// TIA Portal project "OC_test_FFT" (V13)

(* hardware
DEVICE "OpenController"  CPU 1515SP PC
   slot 0: "OpenController"  CPU 1515SP PC  6ES7 677-2AAxx-0xB0  V1.8
      slot 124: "Diagbase"  Diagbase  V6.0.4
      slot 125: "OpenController"  PC Station 2.0  Station_Manager  V2.0
   slot 1: "CPU1505S"  CPU 1505S  6ES7 672-5AC00-0YA0  V1.8
   slot 2: "PROFINET onboard_2"  IE General  IE_CP  V2.0
   slot 4: "HMI_RT_1"  WinCC RT Advanced  6AV2 104-0xxxx-xxxx  13.0.1.0
      slot 33792: "Host interface"  Host interface
   slot 127: "PROFINET BusAdapter CU"  PROFINET Interface  6ES7 193-6AR00-0AA0  V0.0
      slot 32769: "Port_1"  6ES7 193-6AR00-0AA0
      slot 32770: "Port_2"  6ES7 193-6AR00-0AA0
   slot 1002: "Server module_1"  Server module  6ES7 193-6PA00-0AA0  V1.0
      slot 1: "Server module_1"  Server module  6ES7 193-6PA00-0AA0
*)

// ===== PLC "CPU1505S"  CPU 1505S =====

VAR_GLOBAL   // PLC tag table "Default tag table"
   "System_Byte" AT %MB1 : Byte;
   "FirstScan" AT %M1.0 : Bool;
   "DiagStatusUpdate" AT %M1.1 : Bool;
   "AlwaysTRUE" AT %M1.2 : Bool;
   "AlwaysFALSE" AT %M1.3 : Bool;
   "Clock_Byte" AT %MB0 : Byte;
   "Clock_10Hz" AT %M0.0 : Bool;
   "Clock_5Hz" AT %M0.1 : Bool;
   "Clock_2.5Hz" AT %M0.2 : Bool;
   "Clock_2Hz" AT %M0.3 : Bool;
   "Clock_1.25Hz" AT %M0.4 : Bool;
   "Clock_1Hz" AT %M0.5 : Bool;
   "Clock_0.625Hz" AT %M0.6 : Bool;
   "Clock_0.5Hz" AT %M0.7 : Bool;
END_VAR

TYPE "FFT_Filter_RTComplex"
   STRUCT
      re : Real;
      im : Real;
   END_STRUCT;
END_TYPE

DATA_BLOCK "ODK_Params"   // DB1
{ S7_Optimized_Access := 'FALSE' }
VERSION : 0.1
   VAR
      Filter_Load : Struct
      END_STRUCT;
      Filt1 : Struct
      END_STRUCT;
      Filt2 : Struct
      END_STRUCT;
      WaveInput_Load : Struct
      END_STRUCT;
      WaveSetup : Struct
      END_STRUCT;
      GetSamples : Struct
      END_STRUCT;
      WriteSamples : Struct
      END_STRUCT;
   END_VAR
BEGIN
END_DATA_BLOCK

DATA_BLOCK "FFT_Filter_RT_Load_DB"   // DB2
{ S7_Optimized_Access := 'FALSE' }
VERSION : 0.1
// stored: InstanceOfName FFT_Filter_RT_Load
"FFT_Filter_RT_Load"
BEGIN
END_DATA_BLOCK

DATA_BLOCK "FFT_Filter_RTFFT_Filt_DB"   // DB3
{ S7_Optimized_Access := 'FALSE' }
VERSION : 0.1
// stored: InstanceOfName FFT_Filter_RTFFT_Filt
"FFT_Filter_RTFFT_Filt"
BEGIN
END_DATA_BLOCK

DATA_BLOCK "FFT_Filter_RTFFT_Filt_DB_1"   // DB4
{ S7_Optimized_Access := 'FALSE' }
VERSION : 0.1
// stored: InstanceOfName FFT_Filter_RTFFT_Filt
"FFT_Filter_RTFFT_Filt"
BEGIN
END_DATA_BLOCK

DATA_BLOCK "FFT_Filt_Data_Load_DB"   // DB5
{ S7_Optimized_Access := 'FALSE' }
VERSION : 0.1
// stored: InstanceOfName FFT_Filt_Data_Load
"FFT_Filt_Data_Load"
BEGIN
END_DATA_BLOCK

DATA_BLOCK "FFT_Filt_DataWaveSetup_DB"   // DB6
{ S7_Optimized_Access := 'FALSE' }
VERSION : 0.1
// stored: InstanceOfName FFT_Filt_DataWaveSetup
"FFT_Filt_DataWaveSetup"
BEGIN
END_DATA_BLOCK

DATA_BLOCK "FFT_Filt_DataGetSamplesStereo_DB"   // DB7
{ S7_Optimized_Access := 'FALSE' }
VERSION : 0.1
// stored: InstanceOfName FFT_Filt_DataGetSamplesStereo
"FFT_Filt_DataGetSamplesStereo"
BEGIN
END_DATA_BLOCK

DATA_BLOCK "FFT_Filt_DataWriteSamples_DB"   // DB8
{ S7_Optimized_Access := 'FALSE' }
VERSION : 0.1
// stored: InstanceOfName FFT_Filt_DataWriteSamples
"FFT_Filt_DataWriteSamples"
BEGIN
END_DATA_BLOCK

FUNCTION_BLOCK "FFT_Filter_RT_Load"   // FB1, SCL
{ S7_Optimized_Access := 'FALSE' }
VERSION : 0.1
// This block is AUTO GENERATED - DO NOT MODIFY this block!
// Created by ODK_CodeGenerator version 2.0.0.0
// at Sun January 31 20:03:01 2016
// ********************************************************
BEGIN
   //
   // DO NOT CHANGE BELOW OF THIS LINE !!
   // This is an automatic generated block by the
   // ODK_CodeGenerator version 2.0.0.0
   // DO NOT CHANGE !!
   //
   #ODK_Load_Instance(REQ := #REQ,
                      LIBRARY_NAME := #_odk_internal_LIBRARY_NAME,
                      INSTANCE_ID := #_odk_internal_INSTANCE_ID,
                      DONE => #DONE,
                      BUSY => #BUSY,
                      ERROR => #ERROR,
                      STATUS => #STATUS);
   //
   // DO NOT CHANGE !!
   // This is an automatic generated block by the
   // ODK_CodeGenerator version 2.0.0.0
   // DO NOT CHANGE ABOVE OF THIS LINE !!
   //
END_FUNCTION_BLOCK

FUNCTION_BLOCK "FFT_Filter_RT_Unload"   // FB2, SCL
{ S7_Optimized_Access := 'FALSE' }
VERSION : 0.1
// This block is AUTO GENERATED - DO NOT MODIFY this block!
// Created by ODK_CodeGenerator version 2.0.0.0
// at Sun January 31 20:03:01 2016
// ********************************************************
BEGIN
   //
   // DO NOT CHANGE BELOW OF THIS LINE !!
   // This is an automatic generated block by the
   // ODK_CodeGenerator version 2.0.0.0
   // DO NOT CHANGE !!
   //
   #ODK_Unld_Instance(REQ := #REQ,
                      INSTANCE_ID := #_odk_internal_INSTANCE_ID,
                      DONE => #DONE,
                      BUSY => #BUSY,
                      ERROR => #ERROR,
                      STATUS => #STATUS);
   //
   // DO NOT CHANGE !!
   // This is an automatic generated block by the
   // ODK_CodeGenerator version 2.0.0.0
   // DO NOT CHANGE ABOVE OF THIS LINE !!
   //
END_FUNCTION_BLOCK

FUNCTION_BLOCK "FFT_Filter_RTFFT1024p"   // FB3, SCL
{ S7_Optimized_Access := 'FALSE' }
VERSION : 0.1
// This block is AUTO GENERATED - DO NOT MODIFY this block!
// Created by ODK_CodeGenerator version 2.0.0.0
// at Sun January 31 20:03:01 2016
// ********************************************************
BEGIN
   //
   // DO NOT CHANGE BELOW OF THIS LINE !!
   // This is an automatic generated block by the
   // ODK_CodeGenerator version 2.0.0.0
   // DO NOT CHANGE !!
   //
   #_odk_internal_pos := 0;
   FOR #_odk_internal_i := 0 TO 1023 DO
     #_odk_internal_err := WRITE_LITTLE(src_variable := #timeCoef[#_odk_internal_i], dest_array := #_odk_internal_IN_BUFFER, pos := #_odk_internal_pos);
   END_FOR;
   #STATUS := ODK_ExcS(INSTANCE_ID := #_odk_internal_INSTANCE_ID,
                       COMMAND := #_odk_internal_COMMAND,
                       IN_DATA := #_odk_internal_IN_BUFFER,
                       INOUT_DATA := #_odk_internal_tmpDefaultValue,
                       OUT_DATA := #_odk_internal_OUT_BUFFER
   );
   IF #STATUS < 16#7000 THEN
     #_odk_internal_pos := 0;
     FOR #_odk_internal_udt_0 := 0 TO 1023 DO
       #_odk_internal_err := READ_LITTLE(dest_Variable => #freqCoef[#_odk_internal_udt_0].re, src_array := #_odk_internal_OUT_BUFFER, pos := #_odk_internal_pos);
       #_odk_internal_err := READ_LITTLE(dest_Variable => #freqCoef[#_odk_internal_udt_0].im, src_array := #_odk_internal_OUT_BUFFER, pos := #_odk_internal_pos);
     END_FOR;
   END_IF;
   //
   // DO NOT CHANGE !!
   // This is an automatic generated block by the
   // ODK_CodeGenerator version 2.0.0.0
   // DO NOT CHANGE ABOVE OF THIS LINE !!
   //
END_FUNCTION_BLOCK

FUNCTION_BLOCK "FFT_Filter_RTLP_Filter"   // FB4, SCL
{ S7_Optimized_Access := 'FALSE' }
VERSION : 0.1
// This block is AUTO GENERATED - DO NOT MODIFY this block!
// Created by ODK_CodeGenerator version 2.0.0.0
// at Sun January 31 20:03:01 2016
// ********************************************************
BEGIN
   //
   // DO NOT CHANGE BELOW OF THIS LINE !!
   // This is an automatic generated block by the
   // ODK_CodeGenerator version 2.0.0.0
   // DO NOT CHANGE !!
   //
   #_odk_internal_pos := 0;
   FOR #_odk_internal_udt_0 := 0 TO 1023 DO
     #_odk_internal_err := WRITE_LITTLE(src_variable := #freqCoef[#_odk_internal_udt_0].re, dest_array := #_odk_internal_IN_BUFFER, pos := #_odk_internal_pos);
     #_odk_internal_err := WRITE_LITTLE(src_variable := #freqCoef[#_odk_internal_udt_0].im, dest_array := #_odk_internal_IN_BUFFER, pos := #_odk_internal_pos);
   END_FOR;
   #STATUS := ODK_ExcS(INSTANCE_ID := #_odk_internal_INSTANCE_ID,
                       COMMAND := #_odk_internal_COMMAND,
                       IN_DATA := #_odk_internal_IN_BUFFER,
                       INOUT_DATA := #_odk_internal_tmpDefaultValue,
                       OUT_DATA := #_odk_internal_OUT_BUFFER
   );
   IF #STATUS < 16#7000 THEN
     #_odk_internal_pos := 0;
     FOR #_odk_internal_udt_0 := 0 TO 1023 DO
       #_odk_internal_err := READ_LITTLE(dest_Variable => #freqCoefFilt[#_odk_internal_udt_0].re, src_array := #_odk_internal_OUT_BUFFER, pos := #_odk_internal_pos);
       #_odk_internal_err := READ_LITTLE(dest_Variable => #freqCoefFilt[#_odk_internal_udt_0].im, src_array := #_odk_internal_OUT_BUFFER, pos := #_odk_internal_pos);
     END_FOR;
   END_IF;
   //
   // DO NOT CHANGE !!
   // This is an automatic generated block by the
   // ODK_CodeGenerator version 2.0.0.0
   // DO NOT CHANGE ABOVE OF THIS LINE !!
   //
END_FUNCTION_BLOCK

FUNCTION_BLOCK "FFT_Filter_RTIFFT1024p"   // FB5, SCL
{ S7_Optimized_Access := 'FALSE' }
VERSION : 0.1
// This block is AUTO GENERATED - DO NOT MODIFY this block!
// Created by ODK_CodeGenerator version 2.0.0.0
// at Sun January 31 20:03:01 2016
// ********************************************************
BEGIN
   //
   // DO NOT CHANGE BELOW OF THIS LINE !!
   // This is an automatic generated block by the
   // ODK_CodeGenerator version 2.0.0.0
   // DO NOT CHANGE !!
   //
   #_odk_internal_pos := 0;
   FOR #_odk_internal_udt_0 := 0 TO 1023 DO
     #_odk_internal_err := WRITE_LITTLE(src_variable := #freqCoef[#_odk_internal_udt_0].re, dest_array := #_odk_internal_IN_BUFFER, pos := #_odk_internal_pos);
     #_odk_internal_err := WRITE_LITTLE(src_variable := #freqCoef[#_odk_internal_udt_0].im, dest_array := #_odk_internal_IN_BUFFER, pos := #_odk_internal_pos);
   END_FOR;
   #STATUS := ODK_ExcS(INSTANCE_ID := #_odk_internal_INSTANCE_ID,
                       COMMAND := #_odk_internal_COMMAND,
                       IN_DATA := #_odk_internal_IN_BUFFER,
                       INOUT_DATA := #_odk_internal_tmpDefaultValue,
                       OUT_DATA := #_odk_internal_OUT_BUFFER
   );
   IF #STATUS < 16#7000 THEN
     #_odk_internal_pos := 0;
     FOR #_odk_internal_i := 0 TO 1023 DO
       #_odk_internal_err := READ_LITTLE(dest_Variable => #timeCoefOut[#_odk_internal_i], src_array := #_odk_internal_OUT_BUFFER, pos := #_odk_internal_pos);
     END_FOR;
   END_IF;
   //
   // DO NOT CHANGE !!
   // This is an automatic generated block by the
   // ODK_CodeGenerator version 2.0.0.0
   // DO NOT CHANGE ABOVE OF THIS LINE !!
   //
END_FUNCTION_BLOCK

FUNCTION_BLOCK "FFT_Filter_RTFFT_Filt"   // FB6, SCL
{ S7_Optimized_Access := 'FALSE' }
VERSION : 0.1
// This block is AUTO GENERATED - DO NOT MODIFY this block!
// Created by ODK_CodeGenerator version 2.0.0.0
// at Sun January 31 20:03:01 2016
// ********************************************************
BEGIN
   //
   // DO NOT CHANGE BELOW OF THIS LINE !!
   // This is an automatic generated block by the
   // ODK_CodeGenerator version 2.0.0.0
   // DO NOT CHANGE !!
   //
   #_odk_internal_pos := 0;
   FOR #_odk_internal_i := 0 TO 1023 DO
     #_odk_internal_err := WRITE_LITTLE(src_variable := #timeCoef[#_odk_internal_i], dest_array := #_odk_internal_IN_BUFFER, pos := #_odk_internal_pos);
   END_FOR;
   #STATUS := ODK_ExcS(INSTANCE_ID := #_odk_internal_INSTANCE_ID,
                       COMMAND := #_odk_internal_COMMAND,
                       IN_DATA := #_odk_internal_IN_BUFFER,
                       INOUT_DATA := #_odk_internal_tmpDefaultValue,
                       OUT_DATA := #_odk_internal_OUT_BUFFER
   );
   IF #STATUS < 16#7000 THEN
     #_odk_internal_pos := 0;
     FOR #_odk_internal_i := 0 TO 1023 DO
       #_odk_internal_err := READ_LITTLE(dest_Variable => #timeCoefOut[#_odk_internal_i], src_array := #_odk_internal_OUT_BUFFER, pos := #_odk_internal_pos);
     END_FOR;
   END_IF;
   //
   // DO NOT CHANGE !!
   // This is an automatic generated block by the
   // ODK_CodeGenerator version 2.0.0.0
   // DO NOT CHANGE ABOVE OF THIS LINE !!
   //
END_FUNCTION_BLOCK

FUNCTION_BLOCK "FFT_Filt_Data_Load"   // FB7, SCL
{ S7_Optimized_Access := 'FALSE' }
VERSION : 0.1
// This block is AUTO GENERATED - DO NOT MODIFY this block!
// Created by ODK_CodeGenerator version 2.0.0.0
// at Sun January 17 17:54:04 2016
// ********************************************************
BEGIN
   //
   // DO NOT CHANGE BELOW OF THIS LINE !!
   // This is an automatic generated block by the
   // ODK_CodeGenerator version 2.0.0.0
   // DO NOT CHANGE !!
   //
   #ODK_Load_Instance(REQ := #REQ,
                      LIBRARY_NAME := #_odk_internal_LIBRARY_NAME,
                      INSTANCE_ID := #_odk_internal_INSTANCE_ID,
                      DONE => #DONE,
                      BUSY => #BUSY,
                      ERROR => #ERROR,
                      STATUS => #STATUS);
   //
   // DO NOT CHANGE !!
   // This is an automatic generated block by the
   // ODK_CodeGenerator version 2.0.0.0
   // DO NOT CHANGE ABOVE OF THIS LINE !!
   //
END_FUNCTION_BLOCK

FUNCTION_BLOCK "FFT_Filt_Data_Unload"   // FB8, SCL
{ S7_Optimized_Access := 'FALSE' }
VERSION : 0.1
// This block is AUTO GENERATED - DO NOT MODIFY this block!
// Created by ODK_CodeGenerator version 2.0.0.0
// at Sun January 17 17:54:04 2016
// ********************************************************
BEGIN
   //
   // DO NOT CHANGE BELOW OF THIS LINE !!
   // This is an automatic generated block by the
   // ODK_CodeGenerator version 2.0.0.0
   // DO NOT CHANGE !!
   //
   #ODK_Unld_Instance(REQ := #REQ,
                      INSTANCE_ID := #_odk_internal_INSTANCE_ID,
                      DONE => #DONE,
                      BUSY => #BUSY,
                      ERROR => #ERROR,
                      STATUS => #STATUS);
   //
   // DO NOT CHANGE !!
   // This is an automatic generated block by the
   // ODK_CodeGenerator version 2.0.0.0
   // DO NOT CHANGE ABOVE OF THIS LINE !!
   //
END_FUNCTION_BLOCK

FUNCTION_BLOCK "FFT_Filt_DataWaveSetup"   // FB9, SCL
{ S7_Optimized_Access := 'FALSE' }
VERSION : 0.1
// This block is AUTO GENERATED - DO NOT MODIFY this block!
// Created by ODK_CodeGenerator version 2.0.0.0
// at Sun January 17 17:54:04 2016
// ********************************************************
//  Setup file handles for IO operation
BEGIN
   //
   // DO NOT CHANGE BELOW OF THIS LINE !!
   // This is an automatic generated block by the
   // ODK_CodeGenerator version 2.0.0.0
   // DO NOT CHANGE !!
   //
   // Setup file handles for IO operation
   IF NOT #_odk_internal_Last_REQ & #REQ & NOT #BUSY THEN
     #_odk_internal_pos := 0;
     #_odk_internal_tmpStringLen := INT_TO_BYTE(LEN(#inFileName));
     #_odk_internal_IN_BUFFER[#_odk_internal_pos] := BYTE#254;
     #_odk_internal_pos := #_odk_internal_pos + 1;
     #_odk_internal_IN_BUFFER[#_odk_internal_pos] := #_odk_internal_tmpStringLen;
     #_odk_internal_pos := #_odk_internal_pos + 1;
     FOR #_odk_internal_i := 1 TO BYTE_TO_INT(#_odk_internal_tmpStringLen) DO
       #_odk_internal_IN_BUFFER[#_odk_internal_pos] := CHAR_TO_BYTE(#inFileName[#_odk_internal_i]);
       #_odk_internal_pos := #_odk_internal_pos + 1;
     END_FOR;
     #_odk_internal_pos := #_odk_internal_pos + 254 - #_odk_internal_tmpStringLen;
     #_odk_internal_tmpStringLen := INT_TO_BYTE(LEN(#outFileName));
     #_odk_internal_IN_BUFFER[#_odk_internal_pos] := BYTE#254;
     #_odk_internal_pos := #_odk_internal_pos + 1;
     #_odk_internal_IN_BUFFER[#_odk_internal_pos] := #_odk_internal_tmpStringLen;
     #_odk_internal_pos := #_odk_internal_pos + 1;
     FOR #_odk_internal_i := 1 TO BYTE_TO_INT(#_odk_internal_tmpStringLen) DO
       #_odk_internal_IN_BUFFER[#_odk_internal_pos] := CHAR_TO_BYTE(#outFileName[#_odk_internal_i]);
       #_odk_internal_pos := #_odk_internal_pos + 1;
     END_FOR;
     #_odk_internal_pos := #_odk_internal_pos + 254 - #_odk_internal_tmpStringLen;

   END_IF;
   #_odk_internal_Last_REQ := #REQ;
   #ODK_ExcA_Instance(REQ := #REQ,
                      INSTANCE_ID := #_odk_internal_INSTANCE_ID,
                      COMMAND := #_odk_internal_COMMAND,
                      IN_DATA := #_odk_internal_IN_BUFFER,
                      INOUT_DATA := #_odk_internal_tmpDefaultValue,
                      OUT_DATA := #_odk_internal_tmpDefaultValue,
                      DONE => #DONE,
                      BUSY => #BUSY,
                      ERROR => #ERROR,
                      STATUS => #STATUS);
   //
   // DO NOT CHANGE !!
   // This is an automatic generated block by the
   // ODK_CodeGenerator version 2.0.0.0
   // DO NOT CHANGE ABOVE OF THIS LINE !!
   //
END_FUNCTION_BLOCK

FUNCTION_BLOCK "FFT_Filt_DataGetSamplesStereo"   // FB10, SCL
{ S7_Optimized_Access := 'FALSE' }
VERSION : 0.1
// This block is AUTO GENERATED - DO NOT MODIFY this block!
// Created by ODK_CodeGenerator version 2.0.0.0
// at Sun January 17 17:54:04 2016
// ********************************************************
//  Get one filter samlple for processing
BEGIN
   //
   // DO NOT CHANGE BELOW OF THIS LINE !!
   // This is an automatic generated block by the
   // ODK_CodeGenerator version 2.0.0.0
   // DO NOT CHANGE !!
   //
   // Get one filter samlple for processing   
   #_odk_internal_Last_REQ := #REQ;
   #ODK_ExcA_Instance(REQ := #REQ,
                      INSTANCE_ID := #_odk_internal_INSTANCE_ID,
                      COMMAND := #_odk_internal_COMMAND,
                      IN_DATA := #_odk_internal_tmpDefaultValue,
                      INOUT_DATA := #_odk_internal_tmpDefaultValue,
                      OUT_DATA := #_odk_internal_OUT_BUFFER,
                      DONE => #DONE,
                      BUSY => #BUSY,
                      ERROR => #ERROR,
                      STATUS => #STATUS);
   IF NOT #BUSY & #_odk_internal_Last_BUSY & NOT #ERROR THEN
     #_odk_internal_pos := 0;
     FOR #_odk_internal_i := 0 TO 1023 DO
       #_odk_internal_err := READ_LITTLE(dest_Variable => #inputSamplesL[#_odk_internal_i], src_array := #_odk_internal_OUT_BUFFER, pos := #_odk_internal_pos);
     END_FOR;
     FOR #_odk_internal_i := 0 TO 1023 DO
       #_odk_internal_err := READ_LITTLE(dest_Variable => #inputSamplesR[#_odk_internal_i], src_array := #_odk_internal_OUT_BUFFER, pos := #_odk_internal_pos);
     END_FOR;
     #lastSample := BYTE_TO_BOOL(#_odk_internal_OUT_BUFFER[#_odk_internal_pos]);
     #_odk_internal_pos := #_odk_internal_pos + 1;
   END_IF;
   #_odk_internal_Last_BUSY := #BUSY;
   //
   // DO NOT CHANGE !!
   // This is an automatic generated block by the
   // ODK_CodeGenerator version 2.0.0.0
   // DO NOT CHANGE ABOVE OF THIS LINE !!
   //
END_FUNCTION_BLOCK

FUNCTION_BLOCK "FFT_Filt_DataWriteSamples"   // FB11, SCL
{ S7_Optimized_Access := 'FALSE' }
VERSION : 0.1
// This block is AUTO GENERATED - DO NOT MODIFY this block!
// Created by ODK_CodeGenerator version 2.0.0.0
// at Sun January 17 17:54:04 2016
// ********************************************************
//  write processed sample frame into file
BEGIN
   //
   // DO NOT CHANGE BELOW OF THIS LINE !!
   // This is an automatic generated block by the
   // ODK_CodeGenerator version 2.0.0.0
   // DO NOT CHANGE !!
   //
   // write processed sample frame into file
   IF NOT #_odk_internal_Last_REQ & #REQ & NOT #BUSY THEN
     #_odk_internal_pos := 0;
     FOR #_odk_internal_i := 0 TO 1023 DO
       #_odk_internal_err := WRITE_LITTLE(src_variable := #filteredSamplesL[#_odk_internal_i], dest_array := #_odk_internal_IN_BUFFER, pos := #_odk_internal_pos);
     END_FOR;
     FOR #_odk_internal_i := 0 TO 1023 DO
       #_odk_internal_err := WRITE_LITTLE(src_variable := #filteredSamplesR[#_odk_internal_i], dest_array := #_odk_internal_IN_BUFFER, pos := #_odk_internal_pos);
     END_FOR;

   END_IF;
   #_odk_internal_Last_REQ := #REQ;
   #ODK_ExcA_Instance(REQ := #REQ,
                      INSTANCE_ID := #_odk_internal_INSTANCE_ID,
                      COMMAND := #_odk_internal_COMMAND,
                      IN_DATA := #_odk_internal_IN_BUFFER,
                      INOUT_DATA := #_odk_internal_tmpDefaultValue,
                      OUT_DATA := #_odk_internal_tmpDefaultValue,
                      DONE => #DONE,
                      BUSY => #BUSY,
                      ERROR => #ERROR,
                      STATUS => #STATUS);
   //
   // DO NOT CHANGE !!
   // This is an automatic generated block by the
   // ODK_CodeGenerator version 2.0.0.0
   // DO NOT CHANGE ABOVE OF THIS LINE !!
   //
END_FUNCTION_BLOCK

FUNCTION "Filter_Run" : Void   // FC1, FBD
{ S7_Optimized_Access := 'FALSE' }
VERSION : 0.1
BEGIN

REGION Network 1
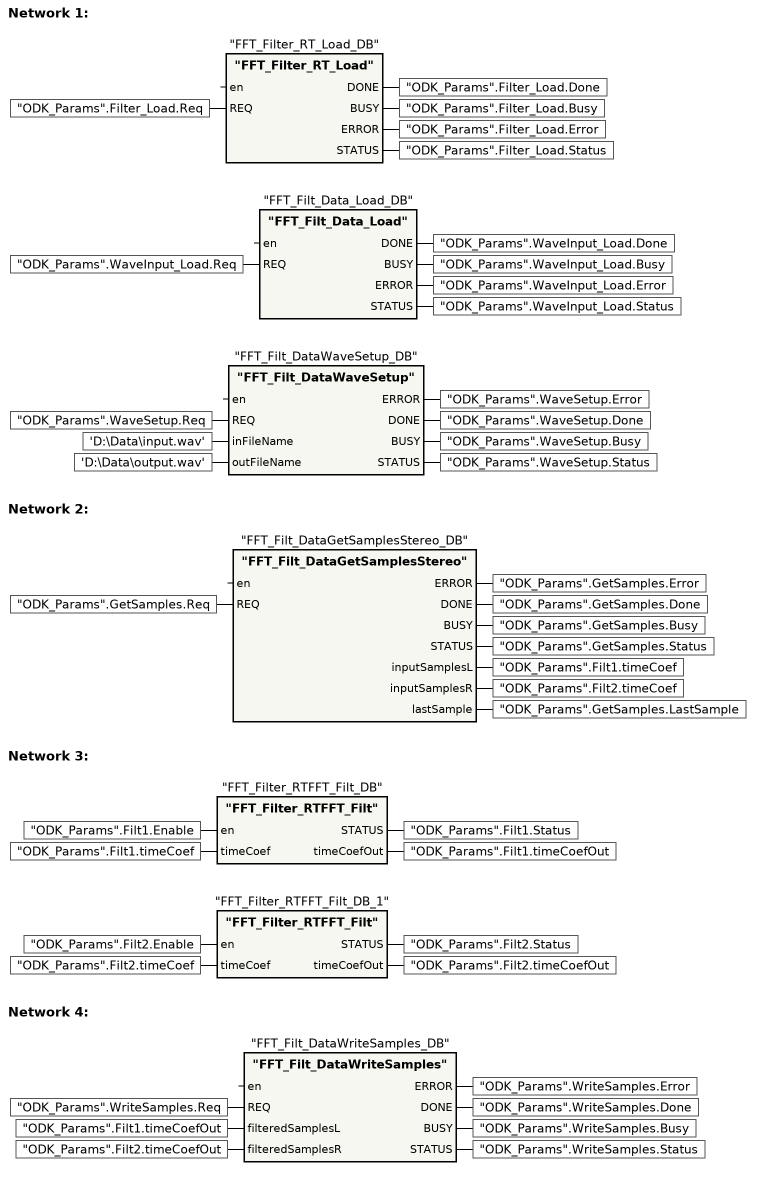
   "FFT_Filter_RT_Load_DB"(REQ := "ODK_Params".Filter_Load.Req,   // "FFT_Filter_RT_Load"
                           DONE => "ODK_Params".Filter_Load.Done,
                           BUSY => "ODK_Params".Filter_Load.Busy,
                           ERROR => "ODK_Params".Filter_Load.Error,
                           STATUS => "ODK_Params".Filter_Load.Status);
   "FFT_Filt_Data_Load_DB"(REQ := "ODK_Params".WaveInput_Load.Req,   // "FFT_Filt_Data_Load"
                           DONE => "ODK_Params".WaveInput_Load.Done,
                           BUSY => "ODK_Params".WaveInput_Load.Busy,
                           ERROR => "ODK_Params".WaveInput_Load.Error,
                           STATUS => "ODK_Params".WaveInput_Load.Status);
   "FFT_Filt_DataWaveSetup_DB"(REQ := "ODK_Params".WaveSetup.Req,   // "FFT_Filt_DataWaveSetup"
                           inFileName := 'D:\Data\input.wav',
                           outFileName := 'D:\Data\output.wav',
                           ERROR => "ODK_Params".WaveSetup.Error,
                           DONE => "ODK_Params".WaveSetup.Done,
                           BUSY => "ODK_Params".WaveSetup.Busy,
                           STATUS => "ODK_Params".WaveSetup.Status);
END_REGION

REGION Network 2
   "FFT_Filt_DataGetSamplesStereo_DB"(REQ := "ODK_Params".GetSamples.Req,   // "FFT_Filt_DataGetSamplesStereo"
                           ERROR => "ODK_Params".GetSamples.Error,
                           DONE => "ODK_Params".GetSamples.Done,
                           BUSY => "ODK_Params".GetSamples.Busy,
                           STATUS => "ODK_Params".GetSamples.Status,
                           inputSamplesL => "ODK_Params".Filt1.timeCoef,
                           inputSamplesR => "ODK_Params".Filt2.timeCoef,
                           lastSample => "ODK_Params".GetSamples.LastSample);
END_REGION

REGION Network 3
   IF "ODK_Params".Filt1.Enable THEN
       "FFT_Filter_RTFFT_Filt_DB"(timeCoef := "ODK_Params".Filt1.timeCoef,   // "FFT_Filter_RTFFT_Filt"
                               STATUS => "ODK_Params".Filt1.Status,
                               timeCoefOut => "ODK_Params".Filt1.timeCoefOut);
   END_IF;
   IF "ODK_Params".Filt2.Enable THEN
       "FFT_Filter_RTFFT_Filt_DB_1"(timeCoef := "ODK_Params".Filt2.timeCoef,   // "FFT_Filter_RTFFT_Filt"
                               STATUS => "ODK_Params".Filt2.Status,
                               timeCoefOut => "ODK_Params".Filt2.timeCoefOut);
   END_IF;
END_REGION

REGION Network 4
   "FFT_Filt_DataWriteSamples_DB"(REQ := "ODK_Params".WriteSamples.Req,   // "FFT_Filt_DataWriteSamples"
                           filteredSamplesL := "ODK_Params".Filt1.timeCoefOut,
                           filteredSamplesR := "ODK_Params".Filt2.timeCoefOut,
                           ERROR => "ODK_Params".WriteSamples.Error,
                           DONE => "ODK_Params".WriteSamples.Done,
                           BUSY => "ODK_Params".WriteSamples.Busy,
                           STATUS => "ODK_Params".WriteSamples.Status);
END_REGION
END_FUNCTION

ORGANIZATION_BLOCK "Main"   // OB1, LAD, ProgramCycle
TITLE = "Main Program Sweep (Cycle)"
{ S7_Optimized_Access := 'FALSE' }
VERSION : 0.1
BEGIN

REGION Network 1
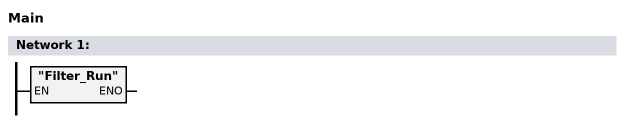
   RUNG wire#powerrail
      "Filter_Run"()
   END_RUNG
   // the same network as SCL:
   "Filter_Run"();
END_REGION
END_ORGANIZATION_BLOCK

(* ===== HMI "HMI_RT_1" =====
connection "HMI_Connection_1": Softbus, S7_1500_OMS

HMI tags "Default tag table"
   "ODK_Params_Filter_Load_Status" : Int, 100 ms
   "ODK_Params_Filter_Load_Req" : Bool, 100 ms
   "ODK_Params_WaveInput_Load_Status" : Int, 100 ms
   "ODK_Params_WaveSetup_Status" : Int, 100 ms
   "ODK_Params_WaveInput_Load_Req" : Bool, 100 ms
   "ODK_Params_WaveSetup_Req" : Bool, 100 ms

screen "Main" 800x600
   TextField "Text field_1" at 50,240 size 112x22
   IOField "I/O field_1" at 62,313 size 93x32
   Button "Button_1" at 62,273 size 96x32
   Button "Button_2" at 62,358 size 96x32
   TextField "Text field_2" at 200,240 size 83x22
   IOField "I/O field_2" at 200,313 size 93x32
   Button "Button_3" at 200,273 size 96x32
   Button "Button_4" at 200,358 size 96x32
   TextField "Text field_3" at 359,240 size 78x22
   IOField "I/O field_3" at 351,313 size 93x32
   Button "Button_5" at 351,273 size 96x32
   Button "Button_6" at 351,358 size 96x32
*)